// TIA Portal project "Delta_Praktika_0" (V17)

(* hardware
DEVICE "S7-1500/ET200MP station_1"  S7-1500 station
   slot 0: "Rail_0"  Rack  6ES7 590-1***0-0AA0
   slot 1: "PLC_2"  CPU 1517TF-3 PN/DP  6ES7 517-3UP00-0AB0  V2.9
      slot 3: "CPU display_1"  6ES7591-1BA00-0AA0
      slot 32768: "PROFINET interface_1"  X1
      slot 33024: "PROFINET interface_2"  X2
      slot 33280: "DP interface_1"  X3
      slot 34817: "Virtual CP interface port_1"  Virtual CP interface port  Virtual CP interface port
DEVICE "ET 200SP station_1"  ET 200SP-Station
   slot 0: "Rack_0"  Rack  6ES5 710-8MAx1
   slot 0: "et200sp"  IM 155-6 PN/2 HF  6ES7 155-6AU01-0CN0  V4.2
   slot 1: "DI 8x24VDC HF_1"  DI 8x24VDC HF  6ES7 131-6BF00-0CA0  V2.0
      slot 1: "DI 8x24VDC HF_1"  DI 8x24VDC HF
   slot 2: "DQ 8x24VDC/0.5A HF_1"  DQ 8x24VDC/0.5A HF  6ES7 132-6BF00-0CA0  V2.0
      slot 1: "DQ 8x24VDC/0.5A HF_1"  DQ 8x24VDC/0.5A HF
   slot 3: "CM 4xIO-Link_1"  CM 4xIO-Link  6ES7 137-6BD00-0BA0  V2.2
      slot 1: "CM 4xIO-Link_1"  6ES7 137-6BD00-0BA0
   slot 4: "Server module_1"  Server module  6ES7 193-6PA00-0AA0  V1.1
      slot 1: "Server module_1"  Server module
   slot 127: "BA 2xRJ45"  BA 2xRJ45  6ES7 193-6AR00-0AA0  V0.0
      slot 1: "Port_1"  X1 P1 R  6ES7 193-6AR00-0AA0  V0.0
      slot 2: "Port_2"  X1 P2 R  6ES7 193-6AR00-0AA0  V0.0
DEVICE "SINAMICS V_1"  SINAMICS V
   slot 0: "SINAMICS V90 PN Rack"  Rail  1.0
   slot 0: "a1"  V90 PN  6SL3 210-5FB10-4UFx  V1.4
      slot 1: "Drive object"  Drive Object
         slot 1: "Module access point"  Module Access Point
         slot 2: "Without PROFIsafe"  No ProfiSafe
         slot 3: "Telegram"  SIEMENS Telegramm 105
DEVICE "SINAMICS V_2"  SINAMICS V
   slot 0: "SINAMICS V90 PN Rack"  Rail  1.0
   slot 0: "a3"  V90 PN  6SL3 210-5FB10-4UFx  V1.4
      slot 1: "Drive object"  Drive Object
         slot 1: "Module access point"  Module Access Point
         slot 2: "Without PROFIsafe"  No ProfiSafe
         slot 3: "Telegram"  SIEMENS Telegramm 105
DEVICE "SINAMICS V_3"  SINAMICS V
   slot 0: "SINAMICS V90 PN Rack"  Rail  1.0
   slot 0: "a2"  V90 PN  6SL3 210-5FB10-4UFx  V1.4
      slot 1: "Drive object"  Drive Object
         slot 1: "Module access point"  Module Access Point
         slot 2: "Without PROFIsafe"  No ProfiSafe
         slot 3: "Telegram"  SIEMENS Telegramm 105
DEVICE "HMI_1"  KTP1200 Basic PN
   slot 0: "HMI_1"  KTP1200 Basic PN  6AV2 123-2MB03-0AX0  17.0.0.0
   slot 1: "HMI_RT_1"  KTP1200 Basic PN  6AV2 123-2MB03-0AX0  17.0.0.0
   slot 5: "HMI_1.IE_CP_1"  PROFINET Interface  17.0.0.0
      slot 1: "Interfaz PROFINET_1"  PROFINET Interface
         slot 1: "Port_1"  Port
*)

// ===== PLC "PLC_2"  CPU 1517TF-3 PN/DP =====
// protected blocks, not shown: "Main_Safety_RTG1", "Main_Safety_RTG1_DB"

VAR_GLOBAL   // PLC tag table "Default tag table"
   "A1_Actor_Interface_AddressIn" AT %I0.0 : "PD_TEL3_IN";
   "A1_Actor_Interface_AddressOut" AT %Q0.0 : "PD_TEL3_OUT";
   "A2_Actor_Interface_AddressIn" AT %I18.0 : "PD_TEL3_IN";
   "A2_Actor_Interface_AddressOut" AT %Q10.0 : "PD_TEL3_OUT";
   "A3_Actor_Interface_AddressIn" AT %I36.0 : "PD_TEL3_IN";
   "A3_Actor_Interface_AddressOut" AT %Q20.0 : "PD_TEL3_OUT";
   "A1_axis_Actor_Interface_AddressIn" AT %I0.0 : "PD_TEL105_IN";
   "A1_axis_Actor_Interface_AddressOut" AT %Q0.0 : "PD_TEL105_OUT";
   "a2_axis_Actor_Interface_AddressIn" AT %I20.0 : "PD_TEL105_IN";
   "a2_axis_Actor_Interface_AddressOut" AT %Q63.0 : "PD_TEL105_OUT";
   "a3_asix_Actor_Interface_AddressIn" AT %I87.0 : "PD_TEL105_IN";
   "a3_asix_Actor_Interface_AddressOut" AT %Q83.0 : "PD_TEL105_OUT";
   "F_Power_Axis1" AT %M20.0 : Bool;
   "F_Power_Axis2" AT %M20.1 : Bool;
   "F_Power_Axis3" AT %M20.2 : Bool;
   "F_Home_Axis1" AT %M20.3 : Bool;
   "F_Home_Axis2" AT %M20.4 : Bool;
   "F_Home_Axis3" AT %M20.5 : Bool;
   "Tag_1" AT %M21.0 : Bool;
   "Tag_2" AT %M21.1 : Bool;
   "Tag_3" AT %M21.2 : Bool;
   "Tag_4" AT %M21.3 : Bool;
   "Tag_5" AT %M21.4 : Bool;
   "Tag_6" AT %M100.0 : Bool;
   "Tag_7" AT %M22.0 : Bool;
   "Tag_8" AT %M22.1 : Bool;
   "Tag_9" AT %M22.2 : Bool;
   "Tag_10" AT %M22.3 : Bool;
   "Tag_11" AT %M22.4 : Bool;
   "Tag_12" AT %M22.5 : Bool;
   "Tag_13" AT %M100.1 : Bool;
   "Tag_14" AT %M22.6 : Bool;
   "Tag_15" AT %Q30.1 : Bool;
   "Tag_16" AT %Q30.0 : Bool;
   "Tag_17" AT %Q30.2 : Bool;
   "Tag_18" AT %M30.1 : Bool;
   "Tag_19" AT %M30.2 : Bool;
   "Tag_20" AT %M30.0 : Bool;
   "Tag_21" AT %M22.7 : Bool;
END_VAR

ORGANIZATION_BLOCK "Main"   // OB1, LAD, ProgramCycle
TITLE = "Main Program Sweep (Cycle)"
{ S7_Optimized_Access := 'TRUE' }
VERSION : 0.1
   VAR_INPUT
      Initial_Call : Bool;   // Initial call of this OB
      Remanence : Bool;   // =True, if remanent data are available
   END_VAR
BEGIN
END_ORGANIZATION_BLOCK

(* ===== HMI "HMI_RT_1" =====
system functions are stored by id; their names below are inferred from use
connection "HMI_Conexión_2": ETHERNET, SMART_S7_1500_OMS

HMI tags "Tabla de variables estándar"
   "F_Power_Axis1" : Bool = PLC F_Power_Axis1 AT %M20.0, 1 s
   "Tag_15" : Bool = PLC Tag_15 AT %Q30.1, 1 s

screen "Imagen_1" 1280x800
   Button "Botón_1" at 38,159 size 96x32; TextOff 'A1+'
   Button "Botón_2" at 175,159 size 96x32; TextOff 'A1-'
   Button "Botón_3" at 40,207 size 96x32; TextOff 'A2+'
   Button "Botón_4" at 175,207 size 96x32; TextOff 'A2-'
   Button "Botón_5" at 40,255 size 96x32; TextOff 'A3+'
   Button "Botón_6" at 175,255 size 96x32; TextOff 'A3-'
   Button "Botón_7" at 308,159 size 96x32; TextOff 'Freno A1'
   Button "Botón_8" at 308,207 size 96x32; TextOff 'Freno A2'
   Button "Botón_9" at 308,255 size 96x32; TextOff 'Freno A3'
   Button "Botón_10" at 926,70 size 96x32; TextOff 'Stop'
   Button "Botón_11" at 1061,70 size 96x32; TextOff 'Reset'
   TextField "Campo de texto_1" at 68,12 size 306x23; Text 'OBJETO TEKNOLOGIKOA BANAKA'
   TextField "Campo de texto_2" at 850,14 size 146x23; Text 'DELTA ROBOTA'
   Circle "Círculo_1" at 415,164 size 19x19
      Appearance <- "Tag_15"
   TextField "Campo de texto_3" at 144,116 size 330x23; Text 'Frenoa desaktibatuta badago berde'
   IOField "Campo ES_1" at 928,418 size 73x30; FormatPattern 99999
   IOField "Campo ES_2" at 928,452 size 73x30; FormatPattern 99999
   IOField "Campo ES_3" at 928,486 size 73x30; FormatPattern 99999
   Button "Botón_15" at 1048,454 size 96x32; TextOff 'GO!'
   TextField "Campo de texto_4" at 928,382 size 270x23; Text 'Mugimendu absoluto linearra'
   TextField "Campo de texto_5" at 1001,418 size 47x23; Text 'X'
   TextField "Campo de texto_6" at 1001,455 size 47x23; Text 'Y'
   TextField "Campo de texto_7" at 1001,492 size 47x23; Text 'Z'
   IOField "Campo ES_4" at 959,607 size 73x30; FormatPattern 99999
   IOField "Campo ES_5" at 959,641 size 73x30; FormatPattern 99999
   IOField "Campo ES_6" at 959,675 size 73x30; FormatPattern 99999
   Button "Botón_16" at 1017,715 size 96x32; TextOff 'GO!'
   TextField "Campo de texto_8" at 959,545 size 288x23; Text 'Mugimendu absoluto zirkularra'
   TextField "Campo de texto_9" at 1032,607 size 47x23; Text 'X'
   TextField "Campo de texto_10" at 1032,644 size 47x23; Text 'Y'
   TextField "Campo de texto_11" at 1032,681 size 47x23; Text 'Z'
   IOField "Campo ES_7" at 1083,608 size 73x30; FormatPattern 99999
   IOField "Campo ES_8" at 1083,642 size 73x30; FormatPattern 99999
   IOField "Campo ES_9" at 1083,676 size 73x30; FormatPattern 99999
   TextField "Campo de texto_12" at 1159,608 size 47x23; Text 'X'
   TextField "Campo de texto_13" at 1159,645 size 47x23; Text 'Y'
   TextField "Campo de texto_14" at 1159,682 size 47x23; Text 'Z'
   TextField "Campo de texto_15" at 928,575 size 135x23; Text 'Nundik pasatu'
   TextField "Campo de texto_16" at 1079,575 size 142x23; Text 'Azken posizioa'
   IOField "Campo ES_13" at 959,607 size 73x30; FormatPattern 99999
   IOField "Campo ES_14" at 959,641 size 73x30; FormatPattern 99999
   IOField "Campo ES_15" at 959,675 size 73x30; FormatPattern 99999
   Button "Botón_18" at 1017,715 size 96x32; TextOff 'GO!'
   TextField "Campo de texto_21" at 959,545 size 288x23; Text 'Mugimendu absoluto zirkularra'
   TextField "Campo de texto_22" at 1032,607 size 47x23; Text 'X'
   TextField "Campo de texto_23" at 1032,644 size 47x23; Text 'Y'
   TextField "Campo de texto_24" at 1032,681 size 47x23; Text 'Z'
   IOField "Campo ES_16" at 1083,608 size 73x30; FormatPattern 99999
   IOField "Campo ES_17" at 1083,642 size 73x30; FormatPattern 99999
   IOField "Campo ES_18" at 1083,676 size 73x30; FormatPattern 99999
   TextField "Campo de texto_25" at 1159,608 size 47x23; Text 'X'
   TextField "Campo de texto_26" at 1159,645 size 47x23; Text 'Y'
   TextField "Campo de texto_27" at 1159,682 size 47x23; Text 'Z'
   TextField "Campo de texto_28" at 928,575 size 135x23; Text 'Nundik pasatu'
   TextField "Campo de texto_29" at 1079,575 size 142x23; Text 'Azken posizioa'
   IOField "Campo ES_10" at 40,390 size 96x32; FormatPattern 9999999
   IOField "Campo ES_11" at 166,388 size 96x32; FormatPattern 9999999
   IOField "Campo ES_12" at 308,388 size 96x32; FormatPattern 9999999
   TextField "Campo de texto_17" at 68,352 size 46x25; Text 'A1'
   TextField "Campo de texto_18" at 198,352 size 46x25; Text 'A2'
   TextField "Campo de texto_19" at 328,352 size 46x25; Text 'A3'
   IOField "Campo ES_19" at 562,418 size 73x30; FormatPattern 99999
   IOField "Campo ES_20" at 562,452 size 73x30; FormatPattern 99999
   IOField "Campo ES_21" at 562,486 size 73x30; FormatPattern 99999
   Button "Botón_17" at 682,454 size 96x32; TextOff 'GO!'
   TextField "Campo de texto_20" at 562,382 size 264x23; Text 'Mugimendu erlatibo linearra'
   TextField "Campo de texto_30" at 635,418 size 47x23; Text 'X'
   TextField "Campo de texto_31" at 635,455 size 47x23; Text 'Y'
   TextField "Campo de texto_32" at 635,492 size 47x23; Text 'Z'
   IOField "Campo ES_22" at 593,607 size 73x30; FormatPattern 99999
   IOField "Campo ES_23" at 593,641 size 73x30; FormatPattern 99999
   IOField "Campo ES_24" at 593,675 size 73x30; FormatPattern 99999
   Button "Botón_19" at 651,715 size 96x32; TextOff 'GO!'
   TextField "Campo de texto_33" at 593,545 size 282x23; Text 'Mugimendu erlatibo zirkularra'
   TextField "Campo de texto_34" at 666,607 size 47x23; Text 'X'
   TextField "Campo de texto_35" at 666,644 size 47x23; Text 'Y'
   TextField "Campo de texto_36" at 666,681 size 47x23; Text 'Z'
   IOField "Campo ES_25" at 717,608 size 73x30; FormatPattern 99999
   IOField "Campo ES_26" at 717,642 size 73x30; FormatPattern 99999
   IOField "Campo ES_27" at 717,676 size 73x30; FormatPattern 99999
   TextField "Campo de texto_37" at 793,608 size 47x23; Text 'X'
   TextField "Campo de texto_38" at 793,645 size 47x23; Text 'Y'
   TextField "Campo de texto_39" at 793,682 size 47x23; Text 'Z'
   TextField "Campo de texto_40" at 562,575 size 135x23; Text 'Nundik pasatu'
   TextField "Campo de texto_41" at 713,575 size 142x23; Text 'Azken posizioa'
   IOField "Campo ES_28" at 593,607 size 73x30; FormatPattern 99999
   IOField "Campo ES_29" at 593,641 size 73x30; FormatPattern 99999
   IOField "Campo ES_30" at 593,675 size 73x30; FormatPattern 99999
   Button "Botón_20" at 651,715 size 96x32; TextOff 'GO!'
   TextField "Campo de texto_43" at 666,607 size 47x23; Text 'X'
   TextField "Campo de texto_44" at 666,644 size 47x23; Text 'Y'
   TextField "Campo de texto_45" at 666,681 size 47x23; Text 'Z'
   IOField "Campo ES_31" at 717,608 size 73x30; FormatPattern 99999
   IOField "Campo ES_32" at 717,642 size 73x30; FormatPattern 99999
   IOField "Campo ES_33" at 717,676 size 73x30; FormatPattern 99999
   TextField "Campo de texto_46" at 793,608 size 47x23; Text 'X'
   TextField "Campo de texto_47" at 793,645 size 47x23; Text 'Y'
   TextField "Campo de texto_48" at 793,682 size 47x23; Text 'Z'
   TextField "Campo de texto_49" at 562,575 size 135x23; Text 'Nundik pasatu'
   TextField "Campo de texto_50" at 713,575 size 142x23; Text 'Azken posizioa'
   TextField "Campo de texto_42" at 581,326 size 254x25; Text 'MUGIMENDU ERLATIBOAK'
   TextField "Campo de texto_51" at 944,326 size 261x25; Text 'MUGIMENDU ABSOLUTOAK'
   IOField "Campo ES_34" at 532,119 size 96x32; FormatPattern 9999999
   IOField "Campo ES_35" at 532,179 size 96x32; FormatPattern 9999999
   IOField "Campo ES_36" at 532,239 size 96x32; FormatPattern 9999999
   TextField "Campo de texto_52" at 635,123 size 46x25; Text 'X'
   TextField "Campo de texto_53" at 633,181 size 46x25; Text 'Y'
   TextField "Campo de texto_54" at 636,239 size 46x25; Text 'Z'
   TextField "Campo de texto_55" at 506,79 size 284x25; Text 'MOMENTUKO X Y Z POSIZIOA'
   TextField "Campo de texto_56" at 14,304 size 448x25; Text 'MOMENTUKO ARDATZEN POSIZIOA GRADUTAN'
   Button "Botón_21" at 888,150 size 298x100; TextOff 'Pick & Place MARTXA'
   Switch "Interruptor_1" at 52,70 size 64x32; CaptionText 'Switch'; TextOff 'OFF'; TextOn 'ON'
      on SwitchOn: SetBit("F_Power_Axis1")
      on SwitchOff: ResetBit("F_Power_Axis1")
   TextField "Campo de texto_57" at 52,45 size 87x25; Text 'Power A1'
   Switch "Interruptor_2" at 187,70 size 64x32; TextOn 'ON'; CaptionText 'Switch'; TextOff 'OFF'
      on SwitchOff: ResetBit("F_Power_Axis1")
      on SwitchOn: SetBit("F_Power_Axis1")
   TextField "Campo de texto_58" at 187,45 size 87x25; Text 'Power A2'
   Switch "Interruptor_3" at 322,70 size 64x32; TextOn 'ON'; CaptionText 'Switch'; TextOff 'OFF'
      on SwitchOff: ResetBit("F_Power_Axis1")
      on SwitchOn: SetBit("F_Power_Axis1")
   TextField "Campo de texto_59" at 322,45 size 87x25; Text 'Power A3'
*)